REGION Network 364
   RUNG wire#powerrail
      Move(in := "EMS".Carrier[68].SDC_OUT.NextCarrierNum, out1 => "Carrier_68_Next_Carrier_Number")
   END_RUNG
   // the same network as SCL:
   "Carrier_68_Next_Carrier_Number" := "EMS".Carrier[68].SDC_OUT.NextCarrierNum;
END_REGION

REGION Network 365
   RUNG wire#powerrail
      Move(in := "EMS".Carrier[68].SDC_OUT.NextStopPos, out1 => "Carrier_68_Next_Stop_Position")
   END_RUNG
   // the same network as SCL:
   "Carrier_68_Next_Stop_Position" := "EMS".Carrier[68].SDC_OUT.NextStopPos;
END_REGION

REGION Network 366
   RUNG wire#powerrail
      Move(in := "EMS".Carrier[68].SDC_OUT.DriveCmdSpeed, out1 => "Carrier_68_Drive_Command_Speed")
   END_RUNG
   // the same network as SCL:
   "Carrier_68_Drive_Command_Speed" := "EMS".Carrier[68].SDC_OUT.DriveCmdSpeed;
END_REGION

REGION Network 367
   RUNG wire#powerrail
      Move(in := "DuplicateCarrierNumber", out1 => "Carrier_68_Duplicate_Carrier_Number")
   END_RUNG
   // the same network as SCL:
   "Carrier_68_Duplicate_Carrier_Number" := "DuplicateCarrierNumber";
END_REGION

REGION Network 368
   RUNG wire#powerrail
      Move(in := "FirstDuplicateCarrierPosition", out1 => "Carrier_68_First_Duplicate_Carrier_Position")
   END_RUNG
   // the same network as SCL:
   "Carrier_68_First_Duplicate_Carrier_Position" := "FirstDuplicateCarrierPosition";
END_REGION

REGION Network 369
   RUNG wire#powerrail
      Move(in := "SecondDuplicateCarrierPosition", out1 => "Carrier_68_Second_Duplicate_Carrier_Position")
   END_RUNG
   // the same network as SCL:
   "Carrier_68_Second_Duplicate_Carrier_Position" := "SecondDuplicateCarrierPosition";
END_REGION

REGION Network 370
   RUNG wire#powerrail
      Contact( "EMS".Carrier[68].SDC_OUT.HeartBeat )
      Coil( "Carrier_68_Heartbeat" )
   END_RUNG
   // the same network as SCL:
   "Carrier_68_Heartbeat" := "EMS".Carrier[68].SDC_OUT.HeartBeat;
END_REGION

REGION Network 371
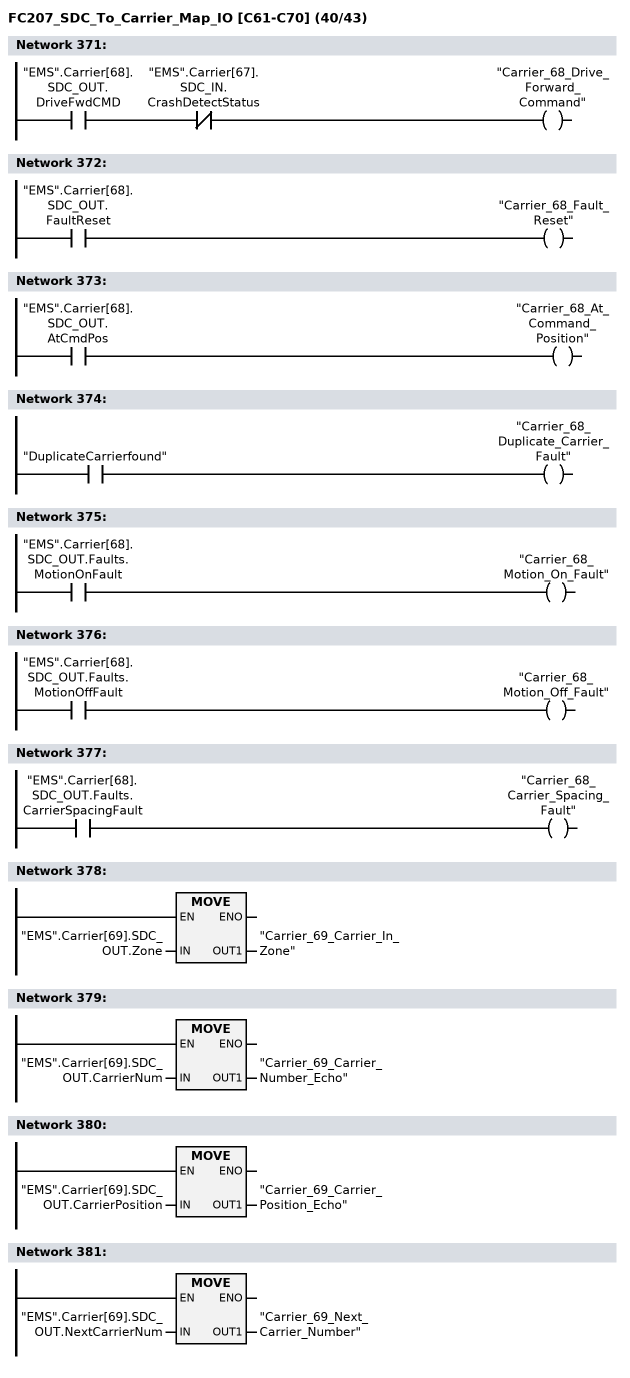
   RUNG wire#powerrail
      Contact( "EMS".Carrier[68].SDC_OUT.DriveFwdCMD )
      I_Contact( "EMS".Carrier[67].SDC_IN.CrashDetectStatus )
      Coil( "Carrier_68_Drive_Forward_Command" )
   END_RUNG
   // the same network as SCL:
   "Carrier_68_Drive_Forward_Command" := "EMS".Carrier[68].SDC_OUT.DriveFwdCMD AND NOT "EMS".Carrier[67].SDC_IN.CrashDetectStatus;
END_REGION

REGION Network 372
   RUNG wire#powerrail
      Contact( "EMS".Carrier[68].SDC_OUT.FaultReset )
      Coil( "Carrier_68_Fault_Reset" )
   END_RUNG
   // the same network as SCL:
   "Carrier_68_Fault_Reset" := "EMS".Carrier[68].SDC_OUT.FaultReset;
END_REGION

REGION Network 373
   RUNG wire#powerrail
      Contact( "EMS".Carrier[68].SDC_OUT.AtCmdPos )
      Coil( "Carrier_68_At_Command_Position" )
   END_RUNG
   // the same network as SCL:
   "Carrier_68_At_Command_Position" := "EMS".Carrier[68].SDC_OUT.AtCmdPos;
END_REGION

REGION Network 374
   RUNG wire#powerrail
      Contact( "DuplicateCarrierfound" )
      Coil( "Carrier_68_Duplicate_Carrier_Fault" )
   END_RUNG
   // the same network as SCL:
   "Carrier_68_Duplicate_Carrier_Fault" := "DuplicateCarrierfound";
END_REGION

REGION Network 375
   RUNG wire#powerrail
      Contact( "EMS".Carrier[68].SDC_OUT.Faults.MotionOnFault )
      Coil( "Carrier_68_Motion_On_Fault" )
   END_RUNG
   // the same network as SCL:
   "Carrier_68_Motion_On_Fault" := "EMS".Carrier[68].SDC_OUT.Faults.MotionOnFault;
END_REGION

REGION Network 376
   RUNG wire#powerrail
      Contact( "EMS".Carrier[68].SDC_OUT.Faults.MotionOffFault )
      Coil( "Carrier_68_Motion_Off_Fault" )
   END_RUNG
   // the same network as SCL:
   "Carrier_68_Motion_Off_Fault" := "EMS".Carrier[68].SDC_OUT.Faults.MotionOffFault;
END_REGION

REGION Network 377
   RUNG wire#powerrail
      Contact( "EMS".Carrier[68].SDC_OUT.Faults.CarrierSpacingFault )
      Coil( "Carrier_68_Carrier_Spacing_Fault" )
   END_RUNG
   // the same network as SCL:
   "Carrier_68_Carrier_Spacing_Fault" := "EMS".Carrier[68].SDC_OUT.Faults.CarrierSpacingFault;
END_REGION

REGION Network 378
   RUNG wire#powerrail
      Move(in := "EMS".Carrier[69].SDC_OUT.Zone, out1 => "Carrier_69_Carrier_In_Zone")
   END_RUNG
   // the same network as SCL:
   "Carrier_69_Carrier_In_Zone" := "EMS".Carrier[69].SDC_OUT.Zone;
END_REGION

REGION Network 379
   RUNG wire#powerrail
      Move(in := "EMS".Carrier[69].SDC_OUT.CarrierNum, out1 => "Carrier_69_Carrier_Number_Echo")
   END_RUNG
   // the same network as SCL:
   "Carrier_69_Carrier_Number_Echo" := "EMS".Carrier[69].SDC_OUT.CarrierNum;
END_REGION

REGION Network 380
   RUNG wire#powerrail
      Move(in := "EMS".Carrier[69].SDC_OUT.CarrierPosition, out1 => "Carrier_69_Carrier_Position_Echo")
   END_RUNG
   // the same network as SCL:
   "Carrier_69_Carrier_Position_Echo" := "EMS".Carrier[69].SDC_OUT.CarrierPosition;
END_REGION

REGION Network 381
   RUNG wire#powerrail
      Move(in := "EMS".Carrier[69].SDC_OUT.NextCarrierNum, out1 => "Carrier_69_Next_Carrier_Number")
   END_RUNG
   // the same network as SCL:
   "Carrier_69_Next_Carrier_Number" := "EMS".Carrier[69].SDC_OUT.NextCarrierNum;
END_REGION

REGION Network 382
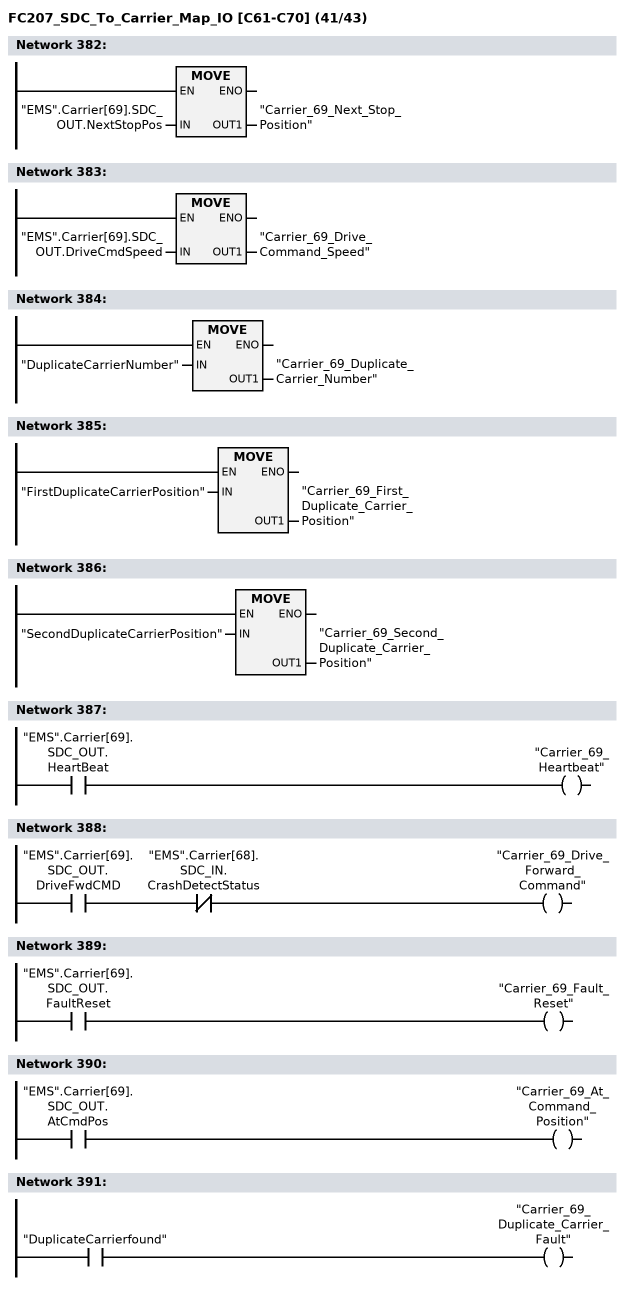
   RUNG wire#powerrail
      Move(in := "EMS".Carrier[69].SDC_OUT.NextStopPos, out1 => "Carrier_69_Next_Stop_Position")
   END_RUNG
   // the same network as SCL:
   "Carrier_69_Next_Stop_Position" := "EMS".Carrier[69].SDC_OUT.NextStopPos;
END_REGION

REGION Network 383
   RUNG wire#powerrail
      Move(in := "EMS".Carrier[69].SDC_OUT.DriveCmdSpeed, out1 => "Carrier_69_Drive_Command_Speed")
   END_RUNG
   // the same network as SCL:
   "Carrier_69_Drive_Command_Speed" := "EMS".Carrier[69].SDC_OUT.DriveCmdSpeed;
END_REGION

REGION Network 384
   RUNG wire#powerrail
      Move(in := "DuplicateCarrierNumber", out1 => "Carrier_69_Duplicate_Carrier_Number")
   END_RUNG
   // the same network as SCL:
   "Carrier_69_Duplicate_Carrier_Number" := "DuplicateCarrierNumber";
END_REGION

REGION Network 385
   RUNG wire#powerrail
      Move(in := "FirstDuplicateCarrierPosition", out1 => "Carrier_69_First_Duplicate_Carrier_Position")
   END_RUNG
   // the same network as SCL:
   "Carrier_69_First_Duplicate_Carrier_Position" := "FirstDuplicateCarrierPosition";
END_REGION

REGION Network 386
   RUNG wire#powerrail
      Move(in := "SecondDuplicateCarrierPosition", out1 => "Carrier_69_Second_Duplicate_Carrier_Position")
   END_RUNG
   // the same network as SCL:
   "Carrier_69_Second_Duplicate_Carrier_Position" := "SecondDuplicateCarrierPosition";
END_REGION

REGION Network 387
   RUNG wire#powerrail
      Contact( "EMS".Carrier[69].SDC_OUT.HeartBeat )
      Coil( "Carrier_69_Heartbeat" )
   END_RUNG
   // the same network as SCL:
   "Carrier_69_Heartbeat" := "EMS".Carrier[69].SDC_OUT.HeartBeat;
END_REGION

REGION Network 388
   RUNG wire#powerrail
      Contact( "EMS".Carrier[69].SDC_OUT.DriveFwdCMD )
      I_Contact( "EMS".Carrier[68].SDC_IN.CrashDetectStatus )
      Coil( "Carrier_69_Drive_Forward_Command" )
   END_RUNG
   // the same network as SCL:
   "Carrier_69_Drive_Forward_Command" := "EMS".Carrier[69].SDC_OUT.DriveFwdCMD AND NOT "EMS".Carrier[68].SDC_IN.CrashDetectStatus;
END_REGION

REGION Network 389
   RUNG wire#powerrail
      Contact( "EMS".Carrier[69].SDC_OUT.FaultReset )
      Coil( "Carrier_69_Fault_Reset" )
   END_RUNG
   // the same network as SCL:
   "Carrier_69_Fault_Reset" := "EMS".Carrier[69].SDC_OUT.FaultReset;
END_REGION

REGION Network 390
   RUNG wire#powerrail
      Contact( "EMS".Carrier[69].SDC_OUT.AtCmdPos )
      Coil( "Carrier_69_At_Command_Position" )
   END_RUNG
   // the same network as SCL:
   "Carrier_69_At_Command_Position" := "EMS".Carrier[69].SDC_OUT.AtCmdPos;
END_REGION

REGION Network 391
   RUNG wire#powerrail
      Contact( "DuplicateCarrierfound" )
      Coil( "Carrier_69_Duplicate_Carrier_Fault" )
   END_RUNG
   // the same network as SCL:
   "Carrier_69_Duplicate_Carrier_Fault" := "DuplicateCarrierfound";
END_REGION

REGION Network 392
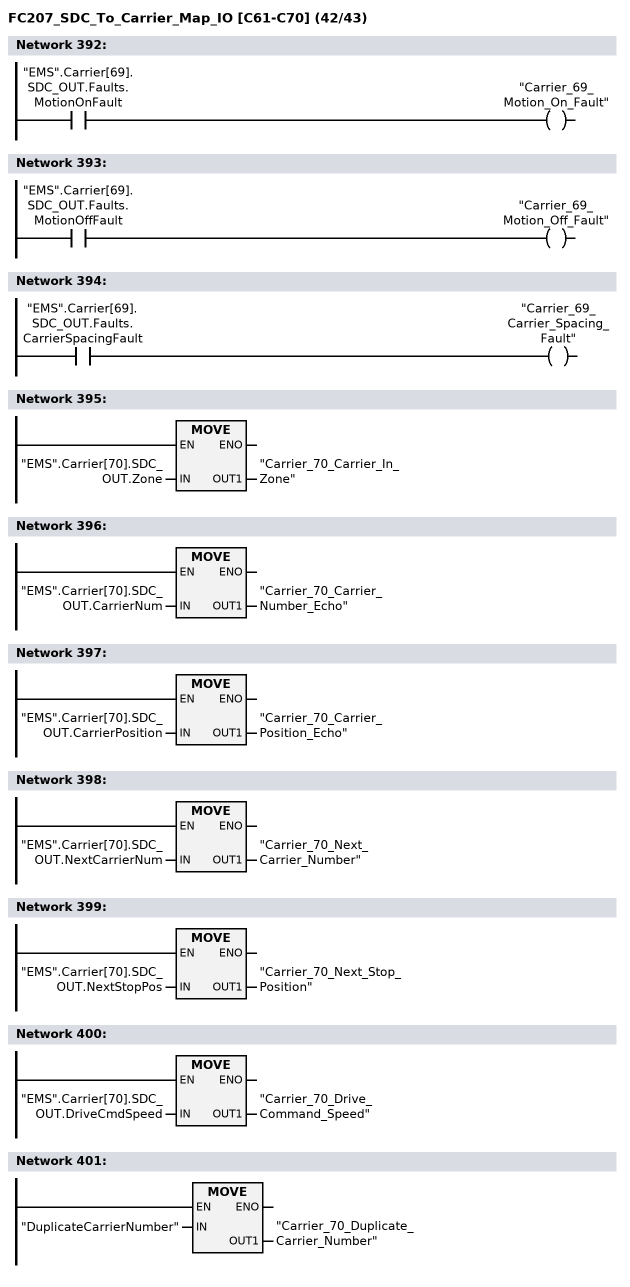
   RUNG wire#powerrail
      Contact( "EMS".Carrier[69].SDC_OUT.Faults.MotionOnFault )
      Coil( "Carrier_69_Motion_On_Fault" )
   END_RUNG
   // the same network as SCL:
   "Carrier_69_Motion_On_Fault" := "EMS".Carrier[69].SDC_OUT.Faults.MotionOnFault;
END_REGION

REGION Network 393
   RUNG wire#powerrail
      Contact( "EMS".Carrier[69].SDC_OUT.Faults.MotionOffFault )
      Coil( "Carrier_69_Motion_Off_Fault" )
   END_RUNG
   // the same network as SCL:
   "Carrier_69_Motion_Off_Fault" := "EMS".Carrier[69].SDC_OUT.Faults.MotionOffFault;
END_REGION

REGION Network 394
   RUNG wire#powerrail
      Contact( "EMS".Carrier[69].SDC_OUT.Faults.CarrierSpacingFault )
      Coil( "Carrier_69_Carrier_Spacing_Fault" )
   END_RUNG
   // the same network as SCL:
   "Carrier_69_Carrier_Spacing_Fault" := "EMS".Carrier[69].SDC_OUT.Faults.CarrierSpacingFault;
END_REGION

REGION Network 395
   RUNG wire#powerrail
      Move(in := "EMS".Carrier[70].SDC_OUT.Zone, out1 => "Carrier_70_Carrier_In_Zone")
   END_RUNG
   // the same network as SCL:
   "Carrier_70_Carrier_In_Zone" := "EMS".Carrier[70].SDC_OUT.Zone;
END_REGION

REGION Network 396
   RUNG wire#powerrail
      Move(in := "EMS".Carrier[70].SDC_OUT.CarrierNum, out1 => "Carrier_70_Carrier_Number_Echo")
   END_RUNG
   // the same network as SCL:
   "Carrier_70_Carrier_Number_Echo" := "EMS".Carrier[70].SDC_OUT.CarrierNum;
END_REGION

REGION Network 397
   RUNG wire#powerrail
      Move(in := "EMS".Carrier[70].SDC_OUT.CarrierPosition, out1 => "Carrier_70_Carrier_Position_Echo")
   END_RUNG
   // the same network as SCL:
   "Carrier_70_Carrier_Position_Echo" := "EMS".Carrier[70].SDC_OUT.CarrierPosition;
END_REGION

REGION Network 398
   RUNG wire#powerrail
      Move(in := "EMS".Carrier[70].SDC_OUT.NextCarrierNum, out1 => "Carrier_70_Next_Carrier_Number")
   END_RUNG
   // the same network as SCL:
   "Carrier_70_Next_Carrier_Number" := "EMS".Carrier[70].SDC_OUT.NextCarrierNum;
END_REGION

REGION Network 399
   RUNG wire#powerrail
      Move(in := "EMS".Carrier[70].SDC_OUT.NextStopPos, out1 => "Carrier_70_Next_Stop_Position")
   END_RUNG
   // the same network as SCL:
   "Carrier_70_Next_Stop_Position" := "EMS".Carrier[70].SDC_OUT.NextStopPos;
END_REGION

REGION Network 400
   RUNG wire#powerrail
      Move(in := "EMS".Carrier[70].SDC_OUT.DriveCmdSpeed, out1 => "Carrier_70_Drive_Command_Speed")
   END_RUNG
   // the same network as SCL:
   "Carrier_70_Drive_Command_Speed" := "EMS".Carrier[70].SDC_OUT.DriveCmdSpeed;
END_REGION

REGION Network 401
   RUNG wire#powerrail
      Move(in := "DuplicateCarrierNumber", out1 => "Carrier_70_Duplicate_Carrier_Number")
   END_RUNG
   // the same network as SCL:
   "Carrier_70_Duplicate_Carrier_Number" := "DuplicateCarrierNumber";
END_REGION

REGION Network 402
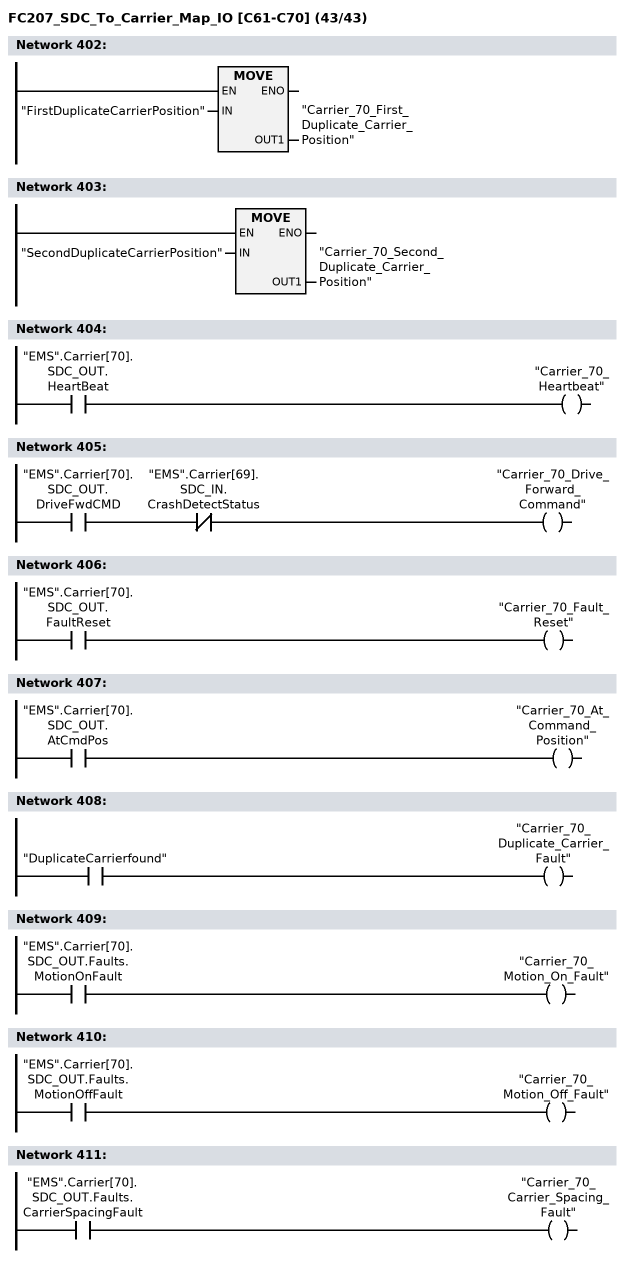
   RUNG wire#powerrail
      Move(in := "FirstDuplicateCarrierPosition", out1 => "Carrier_70_First_Duplicate_Carrier_Position")
   END_RUNG
   // the same network as SCL:
   "Carrier_70_First_Duplicate_Carrier_Position" := "FirstDuplicateCarrierPosition";
END_REGION

REGION Network 403
   RUNG wire#powerrail
      Move(in := "SecondDuplicateCarrierPosition", out1 => "Carrier_70_Second_Duplicate_Carrier_Position")
   END_RUNG
   // the same network as SCL:
   "Carrier_70_Second_Duplicate_Carrier_Position" := "SecondDuplicateCarrierPosition";
END_REGION

REGION Network 404
   RUNG wire#powerrail
      Contact( "EMS".Carrier[70].SDC_OUT.HeartBeat )
      Coil( "Carrier_70_Heartbeat" )
   END_RUNG
   // the same network as SCL:
   "Carrier_70_Heartbeat" := "EMS".Carrier[70].SDC_OUT.HeartBeat;
END_REGION

REGION Network 405
   RUNG wire#powerrail
      Contact( "EMS".Carrier[70].SDC_OUT.DriveFwdCMD )
      I_Contact( "EMS".Carrier[69].SDC_IN.CrashDetectStatus )
      Coil( "Carrier_70_Drive_Forward_Command" )
   END_RUNG
   // the same network as SCL:
   "Carrier_70_Drive_Forward_Command" := "EMS".Carrier[70].SDC_OUT.DriveFwdCMD AND NOT "EMS".Carrier[69].SDC_IN.CrashDetectStatus;
END_REGION

REGION Network 406
   RUNG wire#powerrail
      Contact( "EMS".Carrier[70].SDC_OUT.FaultReset )
      Coil( "Carrier_70_Fault_Reset" )
   END_RUNG
   // the same network as SCL:
   "Carrier_70_Fault_Reset" := "EMS".Carrier[70].SDC_OUT.FaultReset;
END_REGION

REGION Network 407
   RUNG wire#powerrail
      Contact( "EMS".Carrier[70].SDC_OUT.AtCmdPos )
      Coil( "Carrier_70_At_Command_Position" )
   END_RUNG
   // the same network as SCL:
   "Carrier_70_At_Command_Position" := "EMS".Carrier[70].SDC_OUT.AtCmdPos;
END_REGION

REGION Network 408
   RUNG wire#powerrail
      Contact( "DuplicateCarrierfound" )
      Coil( "Carrier_70_Duplicate_Carrier_Fault" )
   END_RUNG
   // the same network as SCL:
   "Carrier_70_Duplicate_Carrier_Fault" := "DuplicateCarrierfound";
END_REGION

REGION Network 409
   RUNG wire#powerrail
      Contact( "EMS".Carrier[70].SDC_OUT.Faults.MotionOnFault )
      Coil( "Carrier_70_Motion_On_Fault" )
   END_RUNG
   // the same network as SCL:
   "Carrier_70_Motion_On_Fault" := "EMS".Carrier[70].SDC_OUT.Faults.MotionOnFault;
END_REGION

REGION Network 410
   RUNG wire#powerrail
      Contact( "EMS".Carrier[70].SDC_OUT.Faults.MotionOffFault )
      Coil( "Carrier_70_Motion_Off_Fault" )
   END_RUNG
   // the same network as SCL:
   "Carrier_70_Motion_Off_Fault" := "EMS".Carrier[70].SDC_OUT.Faults.MotionOffFault;
END_REGION

REGION Network 411
   RUNG wire#powerrail
      Contact( "EMS".Carrier[70].SDC_OUT.Faults.CarrierSpacingFault )
      Coil( "Carrier_70_Carrier_Spacing_Fault" )
   END_RUNG
   // the same network as SCL:
   "Carrier_70_Carrier_Spacing_Fault" := "EMS".Carrier[70].SDC_OUT.Faults.CarrierSpacingFault;
END_REGION
END_FUNCTION

FUNCTION "FC208_SDC_To_Carrier_Map_IO [C71-C80]" : Void   // FC208, LAD
{ S7_Optimized_Access := 'TRUE' }
VERSION : 0.1
BEGIN

REGION Network 1
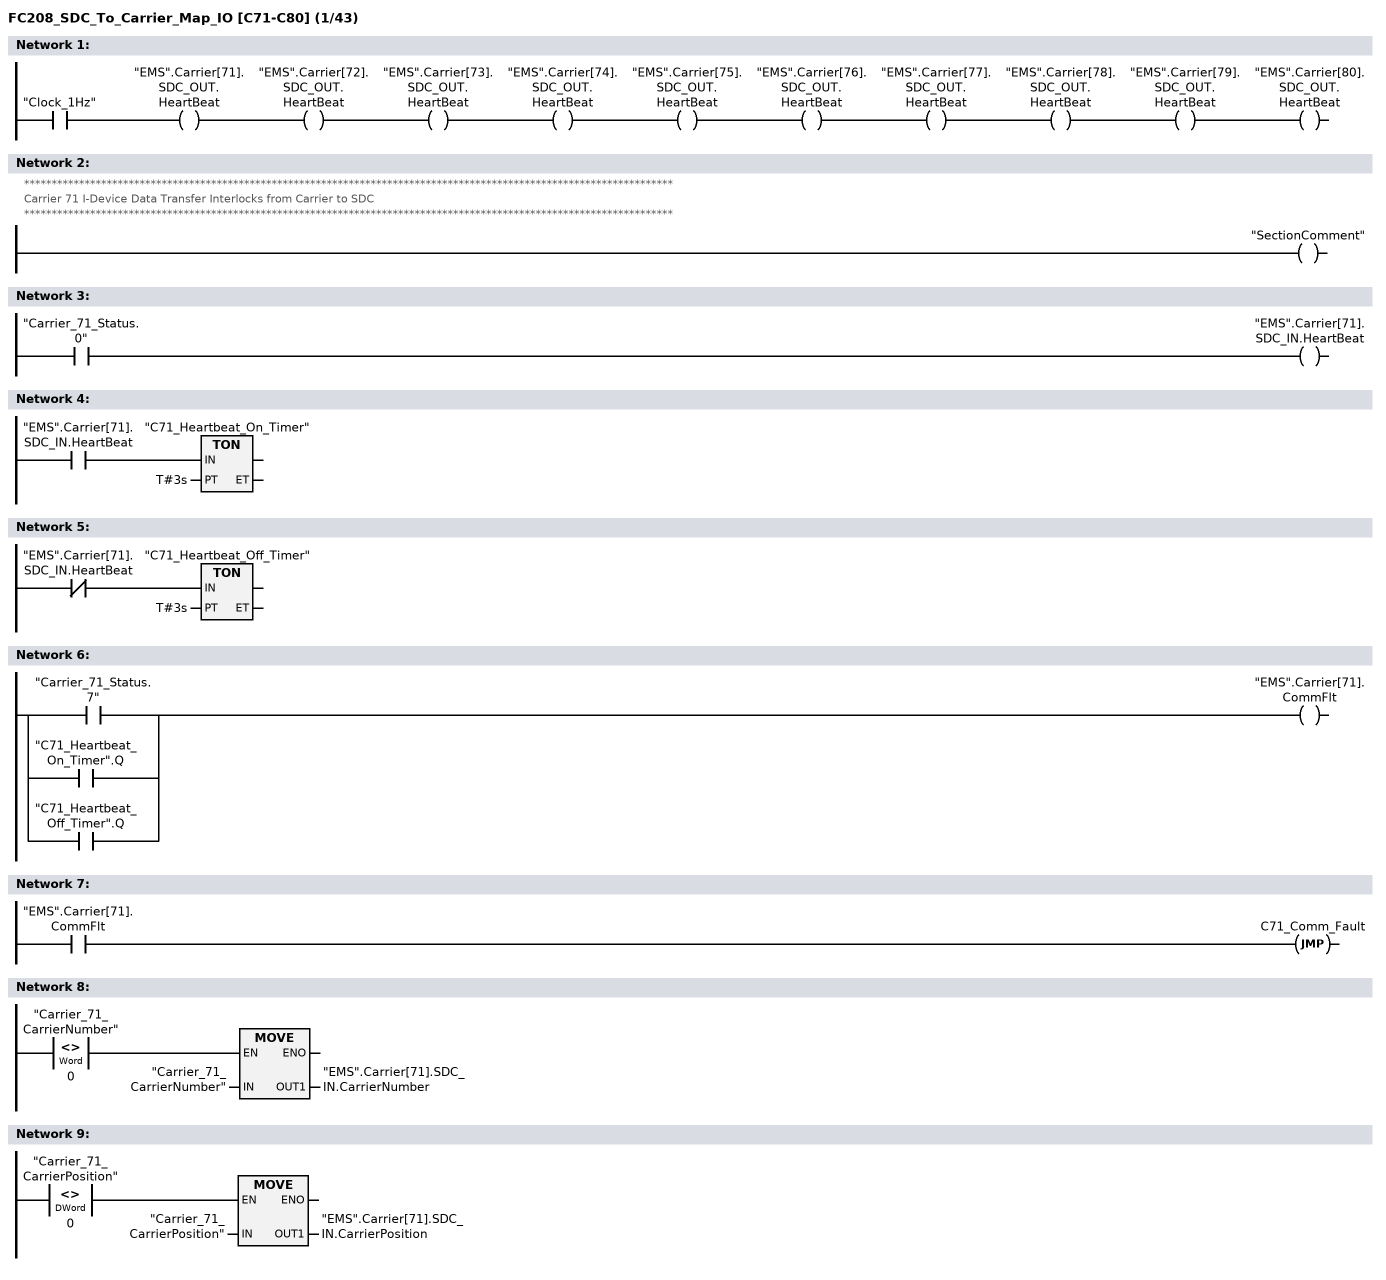
   RUNG wire#powerrail
      Contact( "Clock_1Hz" )
      Coil( "EMS".Carrier[71].SDC_OUT.HeartBeat )
      Coil( "EMS".Carrier[72].SDC_OUT.HeartBeat )
      Coil( "EMS".Carrier[73].SDC_OUT.HeartBeat )
      Coil( "EMS".Carrier[74].SDC_OUT.HeartBeat )
      Coil( "EMS".Carrier[75].SDC_OUT.HeartBeat )
      Coil( "EMS".Carrier[76].SDC_OUT.HeartBeat )
      Coil( "EMS".Carrier[77].SDC_OUT.HeartBeat )
      Coil( "EMS".Carrier[78].SDC_OUT.HeartBeat )
      Coil( "EMS".Carrier[79].SDC_OUT.HeartBeat )
      Coil( "EMS".Carrier[80].SDC_OUT.HeartBeat )
   END_RUNG
   // the same network as SCL:
   "EMS".Carrier[71].SDC_OUT.HeartBeat := "Clock_1Hz";
   "EMS".Carrier[72].SDC_OUT.HeartBeat := "Clock_1Hz";
   "EMS".Carrier[73].SDC_OUT.HeartBeat := "Clock_1Hz";
   "EMS".Carrier[74].SDC_OUT.HeartBeat := "Clock_1Hz";
   "EMS".Carrier[75].SDC_OUT.HeartBeat := "Clock_1Hz";
   "EMS".Carrier[76].SDC_OUT.HeartBeat := "Clock_1Hz";
   "EMS".Carrier[77].SDC_OUT.HeartBeat := "Clock_1Hz";
   "EMS".Carrier[78].SDC_OUT.HeartBeat := "Clock_1Hz";
   "EMS".Carrier[79].SDC_OUT.HeartBeat := "Clock_1Hz";
   "EMS".Carrier[80].SDC_OUT.HeartBeat := "Clock_1Hz";
END_REGION

REGION Network 2
   // **********************************************************************************************************************
   // 
   // Carrier 71 I-Device Data Transfer Interlocks from Carrier to SDC
   // 
   // **********************************************************************************************************************
   RUNG wire#powerrail
      Coil( "SectionComment" )
   END_RUNG
   // the same network as SCL:
   "SectionComment" := TRUE;
END_REGION

REGION Network 3
   RUNG wire#powerrail
      Contact( "Carrier_71_Status.0" )
      Coil( "EMS".Carrier[71].SDC_IN.HeartBeat )
   END_RUNG
   // the same network as SCL:
   "EMS".Carrier[71].SDC_IN.HeartBeat := "Carrier_71_Status.0";
END_REGION

REGION Network 4
   "C71_Heartbeat_On_Timer".TON(IN := "EMS".Carrier[71].SDC_IN.HeartBeat, PT := T#3s);
END_REGION

REGION Network 5
   "C71_Heartbeat_Off_Timer".TON(IN := NOT "EMS".Carrier[71].SDC_IN.HeartBeat, PT := T#3s);
END_REGION

REGION Network 6
   RUNG wire#powerrail
      Contact( "Carrier_71_Status.7" )
      wire#w1
      Coil( "EMS".Carrier[71].CommFlt )
   END_RUNG
   RUNG wire#powerrail
      Contact( "C71_Heartbeat_On_Timer".Q )
   END_RUNG wire#w1
   RUNG wire#powerrail
      Contact( "C71_Heartbeat_Off_Timer".Q )
   END_RUNG wire#w1
   // the same network as SCL:
   "EMS".Carrier[71].CommFlt := "Carrier_71_Status.7" OR "C71_Heartbeat_On_Timer".Q OR "C71_Heartbeat_Off_Timer".Q;
END_REGION

REGION Network 7
   RUNG wire#powerrail
      Contact( "EMS".Carrier[71].CommFlt )
      JumpCoil( C71_Comm_Fault )
   END_RUNG
   // the same network as SCL:
   IF "EMS".Carrier[71].CommFlt THEN GOTO C71_Comm_Fault; END_IF;
END_REGION

REGION Network 8
   RUNG wire#powerrail
      { S7_Templates := "SrcType := Word" } NE_Contact(in1 := "Carrier_71_CarrierNumber", in2 := 0)
      Move(in := "Carrier_71_CarrierNumber", out1 => "EMS".Carrier[71].SDC_IN.CarrierNumber)
   END_RUNG
   // the same network as SCL:
   IF "Carrier_71_CarrierNumber" <> 0 THEN
       "EMS".Carrier[71].SDC_IN.CarrierNumber := "Carrier_71_CarrierNumber";
   END_IF;
END_REGION

REGION Network 9
   RUNG wire#powerrail
      { S7_Templates := "SrcType := DWord" } NE_Contact(in1 := "Carrier_71_CarrierPosition", in2 := 0)
      Move(in := "Carrier_71_CarrierPosition", out1 => "EMS".Carrier[71].SDC_IN.CarrierPosition)
   END_RUNG
   // the same network as SCL:
   IF "Carrier_71_CarrierPosition" <> 0 THEN
       "EMS".Carrier[71].SDC_IN.CarrierPosition := "Carrier_71_CarrierPosition";
   END_IF;
END_REGION

REGION Network 10
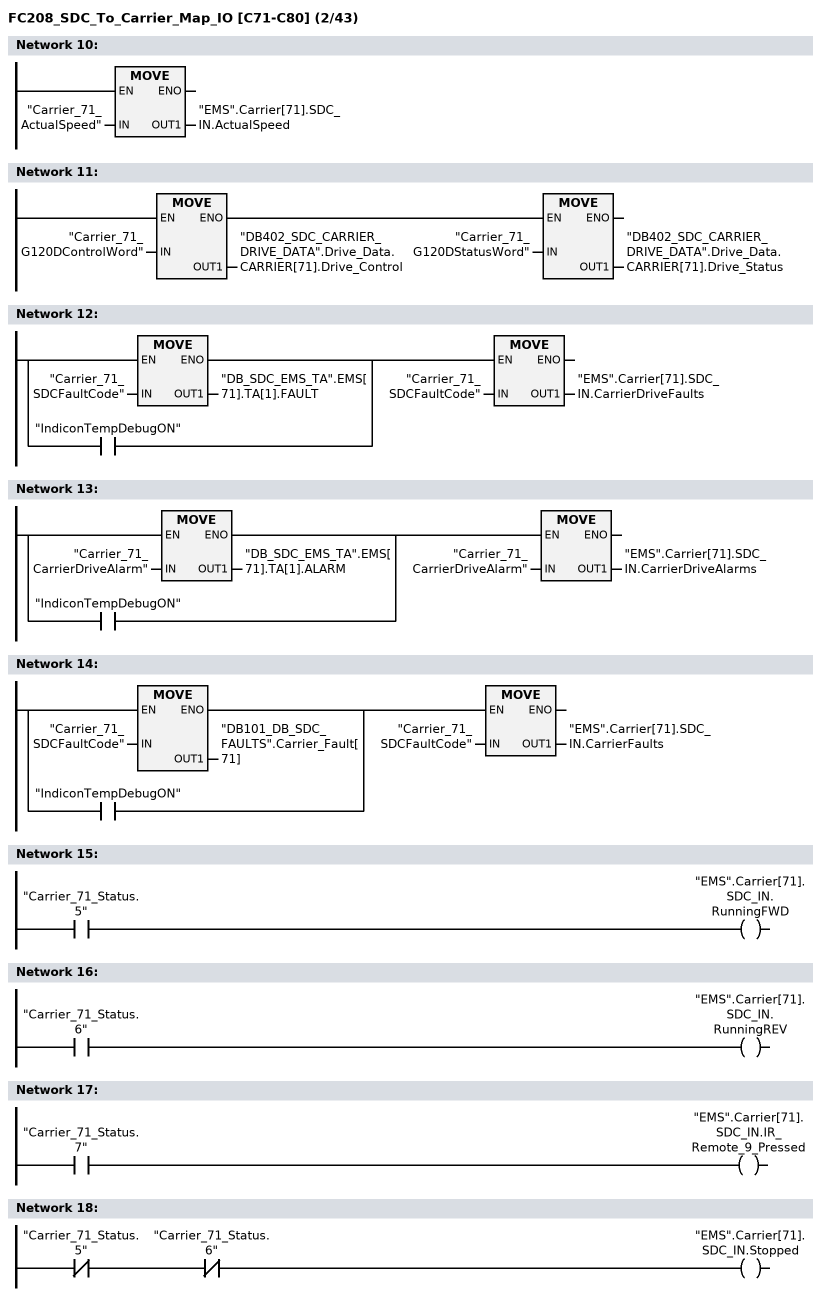
   RUNG wire#powerrail
      Move(in := "Carrier_71_ActualSpeed", out1 => "EMS".Carrier[71].SDC_IN.ActualSpeed)
   END_RUNG
   // the same network as SCL:
   "EMS".Carrier[71].SDC_IN.ActualSpeed := "Carrier_71_ActualSpeed";
END_REGION

REGION Network 11
   RUNG wire#powerrail
      Move(in := "Carrier_71_G120DControlWord", out1 => "DB402_SDC_CARRIER_DRIVE_DATA".Drive_Data.CARRIER[71].Drive_Control)
      Move(in := "Carrier_71_G120DStatusWord", out1 => "DB402_SDC_CARRIER_DRIVE_DATA".Drive_Data.CARRIER[71].Drive_Status)
   END_RUNG
   // the same network as SCL:
   "DB402_SDC_CARRIER_DRIVE_DATA".Drive_Data.CARRIER[71].Drive_Control := "Carrier_71_G120DControlWord";
   "DB402_SDC_CARRIER_DRIVE_DATA".Drive_Data.CARRIER[71].Drive_Status := "Carrier_71_G120DStatusWord";
END_REGION

REGION Network 12
   RUNG wire#powerrail
      Move(in := "Carrier_71_SDCFaultCode", out1 => "DB_SDC_EMS_TA".EMS[71].TA[1].FAULT)
      wire#w1
      Move(in := "Carrier_71_SDCFaultCode", out1 => "EMS".Carrier[71].SDC_IN.CarrierDriveFaults)
   END_RUNG
   RUNG wire#powerrail
      Contact( "IndiconTempDebugON" )
   END_RUNG wire#w1
   // the same network as SCL:
   "DB_SDC_EMS_TA".EMS[71].TA[1].FAULT := "Carrier_71_SDCFaultCode";
   IF TRUE OR "IndiconTempDebugON" THEN
       "EMS".Carrier[71].SDC_IN.CarrierDriveFaults := "Carrier_71_SDCFaultCode";
   END_IF;
END_REGION

REGION Network 13
   RUNG wire#powerrail
      Move(in := "Carrier_71_CarrierDriveAlarm", out1 => "DB_SDC_EMS_TA".EMS[71].TA[1].ALARM)
      wire#w1
      Move(in := "Carrier_71_CarrierDriveAlarm", out1 => "EMS".Carrier[71].SDC_IN.CarrierDriveAlarms)
   END_RUNG
   RUNG wire#powerrail
      Contact( "IndiconTempDebugON" )
   END_RUNG wire#w1
   // the same network as SCL:
   "DB_SDC_EMS_TA".EMS[71].TA[1].ALARM := "Carrier_71_CarrierDriveAlarm";
   IF TRUE OR "IndiconTempDebugON" THEN
       "EMS".Carrier[71].SDC_IN.CarrierDriveAlarms := "Carrier_71_CarrierDriveAlarm";
   END_IF;
END_REGION

REGION Network 14
   RUNG wire#powerrail
      Move(in := "Carrier_71_SDCFaultCode", out1 => "DB101_DB_SDC_FAULTS".Carrier_Fault[71])
      wire#w1
      Move(in := "Carrier_71_SDCFaultCode", out1 => "EMS".Carrier[71].SDC_IN.CarrierFaults)
   END_RUNG
   RUNG wire#powerrail
      Contact( "IndiconTempDebugON" )
   END_RUNG wire#w1
   // the same network as SCL:
   "DB101_DB_SDC_FAULTS".Carrier_Fault[71] := "Carrier_71_SDCFaultCode";
   IF TRUE OR "IndiconTempDebugON" THEN
       "EMS".Carrier[71].SDC_IN.CarrierFaults := "Carrier_71_SDCFaultCode";
   END_IF;
END_REGION

REGION Network 15
   RUNG wire#powerrail
      Contact( "Carrier_71_Status.5" )
      Coil( "EMS".Carrier[71].SDC_IN.RunningFWD )
   END_RUNG
   // the same network as SCL:
   "EMS".Carrier[71].SDC_IN.RunningFWD := "Carrier_71_Status.5";
END_REGION

REGION Network 16
   RUNG wire#powerrail
      Contact( "Carrier_71_Status.6" )
      Coil( "EMS".Carrier[71].SDC_IN.RunningREV )
   END_RUNG
   // the same network as SCL:
   "EMS".Carrier[71].SDC_IN.RunningREV := "Carrier_71_Status.6";
END_REGION

REGION Network 17
   RUNG wire#powerrail
      Contact( "Carrier_71_Status.7" )
      Coil( "EMS".Carrier[71].SDC_IN.IR_Remote_9_Pressed )
   END_RUNG
   // the same network as SCL:
   "EMS".Carrier[71].SDC_IN.IR_Remote_9_Pressed := "Carrier_71_Status.7";
END_REGION

REGION Network 18
   RUNG wire#powerrail
      I_Contact( "Carrier_71_Status.5" )
      I_Contact( "Carrier_71_Status.6" )
      Coil( "EMS".Carrier[71].SDC_IN.Stopped )
   END_RUNG
   // the same network as SCL:
   "EMS".Carrier[71].SDC_IN.Stopped := NOT "Carrier_71_Status.5" AND NOT "Carrier_71_Status.6";
END_REGION

REGION Network 19
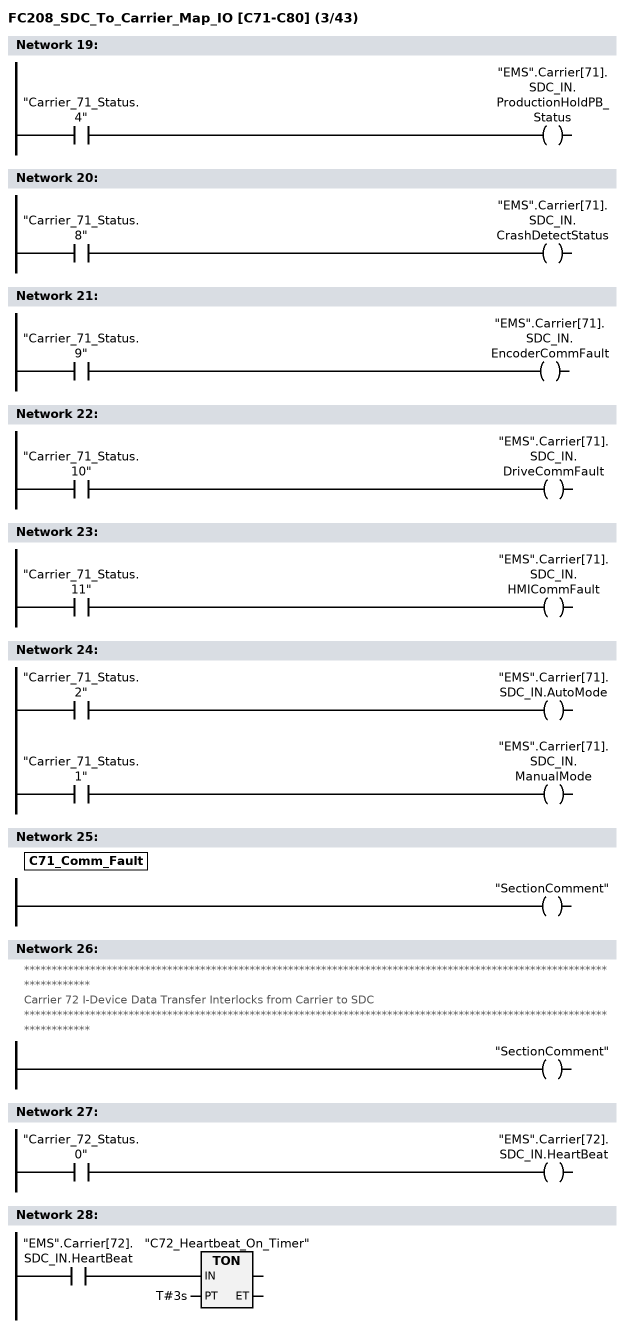
   RUNG wire#powerrail
      Contact( "Carrier_71_Status.4" )
      Coil( "EMS".Carrier[71].SDC_IN.ProductionHoldPB_Status )
   END_RUNG
   // the same network as SCL:
   "EMS".Carrier[71].SDC_IN.ProductionHoldPB_Status := "Carrier_71_Status.4";
END_REGION

REGION Network 20
   RUNG wire#powerrail
      Contact( "Carrier_71_Status.8" )
      Coil( "EMS".Carrier[71].SDC_IN.CrashDetectStatus )
   END_RUNG
   // the same network as SCL:
   "EMS".Carrier[71].SDC_IN.CrashDetectStatus := "Carrier_71_Status.8";
END_REGION

REGION Network 21
   RUNG wire#powerrail
      Contact( "Carrier_71_Status.9" )
      Coil( "EMS".Carrier[71].SDC_IN.EncoderCommFault )
   END_RUNG
   // the same network as SCL:
   "EMS".Carrier[71].SDC_IN.EncoderCommFault := "Carrier_71_Status.9";
END_REGION

REGION Network 22
   RUNG wire#powerrail
      Contact( "Carrier_71_Status.10" )
      Coil( "EMS".Carrier[71].SDC_IN.DriveCommFault )
   END_RUNG
   // the same network as SCL:
   "EMS".Carrier[71].SDC_IN.DriveCommFault := "Carrier_71_Status.10";
END_REGION

REGION Network 23
   RUNG wire#powerrail
      Contact( "Carrier_71_Status.11" )
      Coil( "EMS".Carrier[71].SDC_IN.HMICommFault )
   END_RUNG
   // the same network as SCL:
   "EMS".Carrier[71].SDC_IN.HMICommFault := "Carrier_71_Status.11";
END_REGION

REGION Network 24
   RUNG wire#powerrail
      Contact( "Carrier_71_Status.2" )
      Coil( "EMS".Carrier[71].SDC_IN.AutoMode )
   END_RUNG
   RUNG wire#powerrail
      Contact( "Carrier_71_Status.1" )
      Coil( "EMS".Carrier[71].SDC_IN.ManualMode )
   END_RUNG
   // the same network as SCL:
   "EMS".Carrier[71].SDC_IN.AutoMode := "Carrier_71_Status.2";
   "EMS".Carrier[71].SDC_IN.ManualMode := "Carrier_71_Status.1";
END_REGION

REGION Network 25
   Label( C71_Comm_Fault )
   RUNG wire#powerrail
      Coil( "SectionComment" )
   END_RUNG
   // the same network as SCL:
   C71_Comm_Fault:
   "SectionComment" := TRUE;
END_REGION

REGION Network 26
   // **********************************************************************************************************************
   // 
   // Carrier 72 I-Device Data Transfer Interlocks from Carrier to SDC
   // 
   // **********************************************************************************************************************
   RUNG wire#powerrail
      Coil( "SectionComment" )
   END_RUNG
   // the same network as SCL:
   "SectionComment" := TRUE;
END_REGION

REGION Network 27
   RUNG wire#powerrail
      Contact( "Carrier_72_Status.0" )
      Coil( "EMS".Carrier[72].SDC_IN.HeartBeat )
   END_RUNG
   // the same network as SCL:
   "EMS".Carrier[72].SDC_IN.HeartBeat := "Carrier_72_Status.0";
END_REGION

REGION Network 28
   "C72_Heartbeat_On_Timer".TON(IN := "EMS".Carrier[72].SDC_IN.HeartBeat, PT := T#3s);
END_REGION

REGION Network 29